// TIA Portal project "uppgift2IndustriellIT" (V18)

(* hardware
DEVICE "S7-1500/ET200MP station_1"  S7-1500 station
   slot 0: "Rail_0"  Rack  6ES7 590-1***0-0AA0
   slot 1: "PLC_1"  CPU 1518-4 PN/DP  6ES7 518-4AP00-0AB0  V3.0
      slot 3: "CPU display_1"  6ES7591-1BA00-0AA0
      slot 32768: "PROFINET interface_1"  X1
         slot 32769: "Port_1"  X1 P1
         slot 32770: "Port_2"  X1 P2
      slot 33024: "PROFINET interface_2"  X2
         slot 33025: "Port_1"  X2 P1
      slot 33280: "PROFINET interface GBIT_3"  X3
         slot 33281: "Port_1"  X3 P1
      slot 33536: "DP interface_1"  X4
      slot 34817: "Virtual CP interface port_1"  Virtual CP interface port  Virtual CP interface port
DEVICE "HMI_1"  KTP700 Mobile
   slot 0: "HMI_1"  KTP700 Mobile  6AV2 125-2GB03-0AX0  17.0.0.0
   slot 1: "HMI_RT_1"  KTP700 Mobile  6AV2 125-2GB03-0AX0  17.0.0.0
   slot 5: "HMI_1.IE_CP_1"  PROFINET Interface  17.0.0.0
      slot 1: "PROFINET Interface_1"  PROFINET Interface
         slot 1: "Port_1"  Port
DEVICE "PC-System_1"  SIMATIC PC station
   slot 0: "SIMATIC PC station"  Rail  SIMATIC PC-Station  V1.0
      slot 125: "Stationmanager"  Station_Manager  V6.0.4
   slot 1: "HMI_RT_2"  WinCC RT Advanced  6AV2 104-0xxxx-xxxx  17.0.0.0
      slot 33792: "Computer interface"  Host interface
   slot 2: "IE general_1"  IE General  IE_CP  V8.2.0
      slot 1: "PROFINET interface"  IEGeneral.Interface.8.2.0
*)

// ===== PLC "PLC_1"  CPU 1518-4 PN/DP =====

VAR_GLOBAL   // PLC tag table "Clock/Flanks"
   "Clock_Byte" AT %MB0 : Byte;
   "Clock_10Hz" AT %M0.0 : Bool;
   "Clock_5Hz" AT %M0.1 : Bool;
   "Clock_2.5Hz" AT %M0.2 : Bool;
   "Clock_2Hz" AT %M0.3 : Bool;
   "Clock_1.25Hz" AT %M0.4 : Bool;
   "Clock_1Hz" AT %M0.5 : Bool;
   "Clock_0.625Hz" AT %M0.6 : Bool;
   "Clock_0.5Hz" AT %M0.7 : Bool;
   "PartExitFlank" AT %I3.0 : Bool;
   "CraneExitPosFlank" AT %I3.1 : Bool;
   "HmiEntryFlank" AT %I4.0 : Bool;
   "HmiFlankExit" AT %I4.1 : Bool;
   "FoundToUnloadFlank" AT %I4.2 : Bool;
   "HmiFlankLoad" AT %I5.0 : Bool;
   "HmiFlankUnload" AT %I5.2 : Bool;
   "VisionErrorFlank" AT %I5.4 : Bool;
END_VAR

VAR_GLOBAL   // PLC tag table "FactoryIO"
   "Start Button" AT %I0.0 : Bool;
   "Reset Button" AT %I0.1 : Bool;
   "Stop Button (NC)" AT %I0.2 : Bool;
   "Emergency Stop (NC)" AT %I0.3 : Bool;
   "Part At Entry (NC)" AT %I0.4 : Bool;
   "Part At Load (NC)" AT %I0.5 : Bool;
   "Part At Unload (NC)" AT %I0.6 : Bool;
   "Part At Exit (NC)" AT %I0.7 : Bool;
   "Crane is at Entry-Pos" AT %I1.0 : Bool;
   "Crane is at Exit-Pos" AT %I1.1 : Bool;
   "Crane is at Default-Pos" AT %I1.2 : Bool;
   "Start Light" AT %Q0.0 : Bool;
   "Reset Light" AT %Q0.1 : Bool;
   "Stop Light" AT %Q0.2 : Bool;
   "Protection Stoplight" AT %Q0.3 : Bool;
   "Emitter" AT %Q0.4 : Bool;
   "Signal Tower Green" AT %Q0.5 : Bool;
   "Signal Tower Yellow" AT %Q0.6 : Bool;
   "Signal Tower Red" AT %Q0.7 : Bool;
   "Extend Crane Entry-Side" AT %Q1.0 : Bool;
   "Extend Crane Exit-Side" AT %Q1.1 : Bool;
   "Vision Sensor Entry" AT %IW24 : Int;
   "Crane Current X Position" AT %IW26 : Int;
   "Crane Current Z Position" AT %IW28 : Int;
   "Entry Conveyor" AT %QW20 : Int;
   "Loading Conveyor" AT %QW22 : Int;
   "Unloading Conveyor" AT %QW24 : Int;
   "Set Crane X Position" AT %QW26 : Int;
   "Set Crane Z Position" AT %QW28 : Int;
   "Free Slots in Storage" AT %QW30 : Int;
   "factoryiorunning" AT %I1.3 : Bool;
   "Exit conveyor" AT %QW32 : Int;
   "alarmStuck" AT %QW34 : Int;
   "alarmLoaderFull" AT %QW36 : Int;
   "alarmUnloaderEmpty" AT %QW38 : Int;
END_VAR

// folder: Databases/HmiRelated

DATA_BLOCK "HmiDb"   // DB16
{ S7_Optimized_Access := 'TRUE' }
VERSION : 0.1
   VAR
      HmiOrderMode : Struct
         HmiOrderAmount : Int;
         HmiExecuteOrder : Bool;
         HmiColorSelected : Int;
         HmiPauseOrder : Bool;
         OrderDelivered : Int;
      END_STRUCT;
      ActivateAcutator : Struct
         HmiRunEntryConv : Bool;
         HmiRunExitConv : Bool;
         HmiExtendEntry : Bool;
         HmiExtendExit : Bool;
         HmiRunLoadConv : Bool;
         HmiRunUnloadConv : Bool;
         hmilighttest : Bool;
      END_STRUCT;
      HmiModes : Struct
         ActivateUnloadHmi : Bool;
         HmiStopmode : Bool;
         HmiRunMode : Bool;
         HmiResetMode : Bool;
      END_STRUCT;
      BoxyMover : Int;
      BoxyMover2 : Int;
      ClearStock : Bool;
      ClearCounter : Bool;
      HmiSaveArmCalX : Bool;
      HmiSaveArmCalY : Bool;
      XListColumn : Int;
      YListColumn : Int;
      CalInputVal : Int;
      CurrentPositionX : Int;
      CurrentPositionY : Int;
      oke : String := 'yes';
   END_VAR
BEGIN
END_DATA_BLOCK

DATA_BLOCK "jogmodeDB"   // DB18
{ S7_Optimized_Access := 'TRUE' }
VERSION : 0.1
   VAR
      CraneXjog : Int;
      CraneYjog : Int;
   END_VAR
BEGIN
END_DATA_BLOCK

// folder: Databases/SCLdb

DATA_BLOCK "PositionArray"   // DB9
{ S7_Optimized_Access := 'TRUE' }
VERSION : 0.1
   VAR RETAIN
      YposCraneMM : Array[0..5] of Int;
      XposCraneMM : Array[0..8] of Int;
   END_VAR
BEGIN
   YposCraneMM[0] := 380;
   YposCraneMM[1] := 1540;
   YposCraneMM[2] := 2680;
   YposCraneMM[3] := 3820;
   YposCraneMM[4] := 4950;
   YposCraneMM[5] := 6000;
   XposCraneMM[0] := 1490;
   XposCraneMM[1] := 2635;
   XposCraneMM[2] := 3750;
   XposCraneMM[3] := 4860;
   XposCraneMM[4] := 6000;
   XposCraneMM[5] := 7145;
   XposCraneMM[6] := 8260;
   XposCraneMM[7] := 9380;
   XposCraneMM[8] := 10500;
END_DATA_BLOCK

DATA_BLOCK "PositionUnload_DB"   // DB10
{ S7_Optimized_Access := 'TRUE' }
VERSION : 0.1
// stored: InstanceOfName PositionUnload
"PositionUnload"
BEGIN
END_DATA_BLOCK

DATA_BLOCK "AlreadyFilledSlotArray"   // DB11
{ S7_Optimized_Access := 'TRUE' }
VERSION : 0.1
   VAR RETAIN
      Row1Y : Array[0..5] of Int;   // siffran i array namnet indikterar X axeln: T.ex. Row3Y visar om column 3 är fylld med lådor och index siffran i arrayn indikerar vilken våning i columen som är fylld
      Row2Y : Array[0..5] of Int;
      Row3Y : Array[0..5] of Int;
      Row4Y : Array[0..5] of Int;
      Row5Y : Array[0..5] of Int;
      Row6Y : Array[0..5] of Int;
      Row7Y : Array[0..5] of Int;
      Row8Y : Array[0..5] of Int;
      Row9Y : Array[0..5] of Int;
   END_VAR
BEGIN
   Row4Y[5] := 0;
   Row4Y[4] := 0;
   Row4Y[3] := 0;
   Row4Y[2] := 0;
   Row4Y[1] := 0;
   Row4Y[0] := 0;
   Row3Y[0] := 0;
   Row3Y[1] := 0;
   Row3Y[2] := 0;
   Row3Y[3] := 0;
   Row3Y[4] := 0;
   Row3Y[5] := 0;
   Row2Y[5] := 0;
   Row2Y[4] := 0;
   Row2Y[3] := 0;
   Row2Y[2] := 0;
   Row2Y[1] := 0;
   Row2Y[0] := 0;
   Row8Y[5] := 0;
   Row8Y[4] := 0;
   Row8Y[3] := 0;
   Row8Y[2] := 0;
   Row8Y[1] := 0;
   Row8Y[0] := 0;
   Row7Y[5] := 0;
   Row7Y[4] := 0;
   Row1Y[5] := 0;
   Row1Y[4] := 0;
   Row1Y[3] := 0;
   Row1Y[2] := 0;
   Row1Y[1] := 0;
   Row1Y[0] := 0;
   Row9Y[5] := 0;
   Row9Y[4] := 0;
   Row9Y[3] := 0;
   Row9Y[2] := 0;
   Row9Y[1] := 0;
   Row9Y[0] := 0;
   Row5Y[5] := 0;
   Row5Y[4] := 0;
   Row5Y[3] := 0;
   Row5Y[2] := 0;
   Row5Y[1] := 0;
   Row5Y[0] := 0;
   Row6Y[5] := 0;
   Row6Y[4] := 0;
   Row6Y[3] := 0;
   Row6Y[2] := 0;
   Row6Y[1] := 0;
   Row6Y[0] := 0;
   Row7Y[3] := 0;
   Row7Y[2] := 0;
   Row7Y[1] := 0;
   Row7Y[0] := 0;
END_DATA_BLOCK

DATA_BLOCK "PositionsLOAD_DB"   // DB13
{ S7_Optimized_Access := 'TRUE' }
VERSION : 0.1
// stored: InstanceOfName PositionsLoad
"PositionsLoad"
BEGIN
END_DATA_BLOCK

DATA_BLOCK "resetFill_DB"   // DB21
{ S7_Optimized_Access := 'TRUE' }
VERSION : 0.1
// stored: InstanceOfName resetFill
"resetFill"
BEGIN
END_DATA_BLOCK

// folder: Databases/input/outputDB

DATA_BLOCK "InputsDB"   // DB1
{ S7_Optimized_Access := 'TRUE' }
VERSION : 0.1
   VAR RETAIN
      ConvertedConveyors : Struct
         EntryConvSensorVal : Int := 7500;
         LoadingConvSensorVal : Int := 7500;
         EntryConvScalex : Real;
         LoadingConvScalex : Real;
         ExitConvSensorVal : Int := 7500;
         ExitConvScaleX : Real;
         UnloadingScaleX : Real;
         UnloadingSensorVal : Int := 7500;
      END_STRUCT;
   END_VAR
   VAR
      ConveyorSaveCalVal : Struct
         Normxconverter : Real;
         Save : Bool;
         "DisplayMm/s" : Real;
         Min : Struct
            EntryMin : Int;
            ExitMin : Int;
            LoadMin : Int;
            UnloadMin : Int;
            HmiDisplayMin : Int;
            ActualdisplayMin : Int;
         END_STRUCT;
         Max : Struct
            EntryMax : Int;
            ExitMax : Int;
            LoadMax : Int;
            UnloadMax : Int;
            HmiDisplayMax : Int;
            ActualdisplayMax : Int;
         END_STRUCT;
      END_STRUCT;
      RunConveyor : Struct
         RunEntryConveyor : Bool;
         RunLoadingConveyor : Bool;
         RunUnloadingConveyor : Bool;
         RunExitConveyor : Bool;
      END_STRUCT;
      Crane : Struct
         X : Struct
            XSensorValueNormx : Real;
            XSensorValueScaleX : Int;
            SaveX : Int;
         END_STRUCT;
         Y : Struct
            YSensorValueNormx : Real;
            YSensorValueScalex : Int;
            SaveY : Int;
         END_STRUCT;
         RunArmX : Bool;
         RunArmY : Bool;
      END_STRUCT;
      Sensors : Struct
         "Part Entry" : Bool;
         "Part Load" : Bool;
         "Part Unload" : Bool;
         "Part Exit" : Bool;
         "Crane Entry" : Bool;
         "Crane Exit" : Bool;
         "Crane Default" : Bool;
         "Color Sensor" : Int;
      END_STRUCT;
      Conditions : Struct
         ProtectedStop : Bool;
         HasBeenJogging : Bool;
         VisionError : Bool;
      END_STRUCT;
      FreeSlotCounter : Int := 54;
      ErrorStuck : Bool;
      ConveyorCalibrationPicker : Int := 10;   // Slidern i hmin
      ConveyorCalibrationBarSlider : Int := 7500;
      ConveyorCalibrationBarSliderTEMP : Int;
      YisMoving : Bool;
      XisMoving : Bool;   // Används endast för hmin just nu
      Math200 : Int := 200;
      Math10 : Int;
      AdjustX : Int;
      AdjustY : Int;
      PressAdjustX : Bool;
      PressAdjustY : Bool;
      totalcounter : Int;
      totalremovedcounter : Int;
   END_VAR
BEGIN
END_DATA_BLOCK

DATA_BLOCK "OutputsDB"   // DB2
{ S7_Optimized_Access := 'TRUE' }
VERSION : 0.1
   VAR
      CraneOutput : Struct
         Xmm : Int;
         Xnormx : Real;
         XScalex : Int;
         Ymm : Int;
         Ynormx : Real;
         YScalex : Int;
      END_STRUCT;
      ForkController : Struct
         MoveForkExitLoad : Bool;
         MoveForkEntryLoad : Bool;
         SafetyStopExitUnload : Bool;
      END_STRUCT;
   END_VAR
BEGIN
END_DATA_BLOCK

DATA_BLOCK "Modes"   // DB3
{ S7_Optimized_Access := 'TRUE' }
VERSION : 0.1
   VAR
      Modes : Struct
         RunMode : Bool;
         ResetMode : Bool;
         Unloadmode : Bool;
         RunUnloadConveyor : Bool;
         StoppestMode : Bool;
         JogMode : Bool;
         OrderMode : Bool;
      END_STRUCT;
      Sequences : Struct
         SequenceLoader : Int := 10;
         SequenceUnloader : Int := 10;
         ResetModeSequence : Int := 10;
         SafetyStopSequence : Int := 10;
      END_STRUCT;
      StopMethods : Struct
         SafetyStop : Bool;
         ProductionStop : Bool := true;
      END_STRUCT;
   END_VAR
BEGIN
END_DATA_BLOCK

DATA_BLOCK "ColorDB"   // DB5
{ S7_Optimized_Access := 'TRUE' }
VERSION : 0.1
   VAR
      Gray : Int;
      Green : Int;
      Blue : Int;
      isGray : Int := 1;
      isBlue : Int := 2;
      isGreen : Int := 3;
   END_VAR
BEGIN
END_DATA_BLOCK

// folder: System blocks/Program resources

DATA_BLOCK "ResetWaiterTimer"   // DB4
{ S7_Optimized_Access := 'TRUE' }
AUTHOR : Simatic
FAMILY : IEC
NAME : IEC_TMR
VERSION : 1.0
// stored: InstanceOfName IEC_TIMER
"IEC_TIMER"
BEGIN
END_DATA_BLOCK

DATA_BLOCK "ColorCounter1"   // DB6
{ S7_Optimized_Access := 'TRUE' }
AUTHOR : Simatic
FAMILY : IEC
NAME : CNTR
VERSION : 1.0
// stored: InstanceOfName IEC_COUNTER
"IEC_COUNTER"
BEGIN
END_DATA_BLOCK

DATA_BLOCK "ColorCouter2"   // DB7
{ S7_Optimized_Access := 'TRUE' }
AUTHOR : Simatic
FAMILY : IEC
NAME : CNTR
VERSION : 1.0
// stored: InstanceOfName IEC_COUNTER
"IEC_COUNTER"
BEGIN
END_DATA_BLOCK

DATA_BLOCK "ColorCounter3"   // DB8
{ S7_Optimized_Access := 'TRUE' }
AUTHOR : Simatic
FAMILY : IEC
NAME : CNTR
VERSION : 1.0
// stored: InstanceOfName IEC_COUNTER
"IEC_COUNTER"
BEGIN
END_DATA_BLOCK

DATA_BLOCK "SclDelay"   // DB12
{ S7_Optimized_Access := 'TRUE' }
AUTHOR : Simatic
FAMILY : IEC
NAME : IEC_TMR
VERSION : 1.0
// stored: InstanceOfName IEC_TIMER
"IEC_TIMER"
BEGIN
END_DATA_BLOCK

DATA_BLOCK "SclDelay2"   // DB14
{ S7_Optimized_Access := 'TRUE' }
AUTHOR : Simatic
FAMILY : IEC
NAME : IEC_TMR
VERSION : 1.0
// stored: InstanceOfName IEC_TIMER
"IEC_TIMER"
BEGIN
END_DATA_BLOCK

DATA_BLOCK "ForkWaiter"   // DB15
{ S7_Optimized_Access := 'TRUE' }
AUTHOR : Simatic
FAMILY : IEC
NAME : IEC_TMR
VERSION : 1.0
// stored: InstanceOfName IEC_TIMER
"IEC_TIMER"
BEGIN
END_DATA_BLOCK

DATA_BLOCK "StuckTimer"   // DB17
{ S7_Optimized_Access := 'TRUE' }
AUTHOR : Simatic
FAMILY : IEC
NAME : IEC_TMR
VERSION : 1.0
// stored: InstanceOfName IEC_TIMER
"IEC_TIMER"
BEGIN
END_DATA_BLOCK

DATA_BLOCK "FreeSlotCounter"   // DB19
{ S7_Optimized_Access := 'TRUE' }
AUTHOR : Simatic
FAMILY : IEC
NAME : CNTR
VERSION : 1.0
// stored: InstanceOfName IEC_COUNTER
"IEC_COUNTER"
BEGIN
   CV := 54;
END_DATA_BLOCK

DATA_BLOCK "OrderDeliverCounter"   // DB20
{ S7_Optimized_Access := 'TRUE' }
AUTHOR : Simatic
FAMILY : IEC
NAME : CNTR
VERSION : 1.0
// stored: InstanceOfName IEC_COUNTER
"IEC_COUNTER"
BEGIN
END_DATA_BLOCK

DATA_BLOCK "totalcounter"   // DB22
{ S7_Optimized_Access := 'TRUE' }
AUTHOR : Simatic
FAMILY : IEC
NAME : CNTR
VERSION : 1.0
// stored: InstanceOfName IEC_COUNTER
"IEC_COUNTER"
BEGIN
END_DATA_BLOCK

DATA_BLOCK "totalcounterremoved"   // DB23
{ S7_Optimized_Access := 'TRUE' }
AUTHOR : Simatic
FAMILY : IEC
NAME : CNTR
VERSION : 1.0
// stored: InstanceOfName IEC_COUNTER
"IEC_COUNTER"
BEGIN
END_DATA_BLOCK

DATA_BLOCK "ResetWaiterTimer2"   // DB24
{ S7_Optimized_Access := 'TRUE' }
AUTHOR : Simatic
FAMILY : IEC
NAME : IEC_TMR
VERSION : 1.0
// stored: InstanceOfName IEC_TIMER
"IEC_TIMER"
BEGIN
END_DATA_BLOCK

DATA_BLOCK "waittimer3"   // DB25
{ S7_Optimized_Access := 'TRUE' }
AUTHOR : Simatic
FAMILY : IEC
NAME : IEC_TMR
VERSION : 1.0
// stored: InstanceOfName IEC_TIMER
"IEC_TIMER"
BEGIN
END_DATA_BLOCK

// folder: (top level)

ORGANIZATION_BLOCK "Main"   // OB1, LAD, ProgramCycle
TITLE = "Main Program Sweep (Cycle)"
{ S7_Optimized_Access := 'TRUE' }
VERSION : 0.1
   VAR_INPUT
      Initial_Call : Bool;   // Initial call of this OB
      Remanence : Bool;   // =True, if remanent data are available
   END_VAR
BEGIN

REGION Network 1
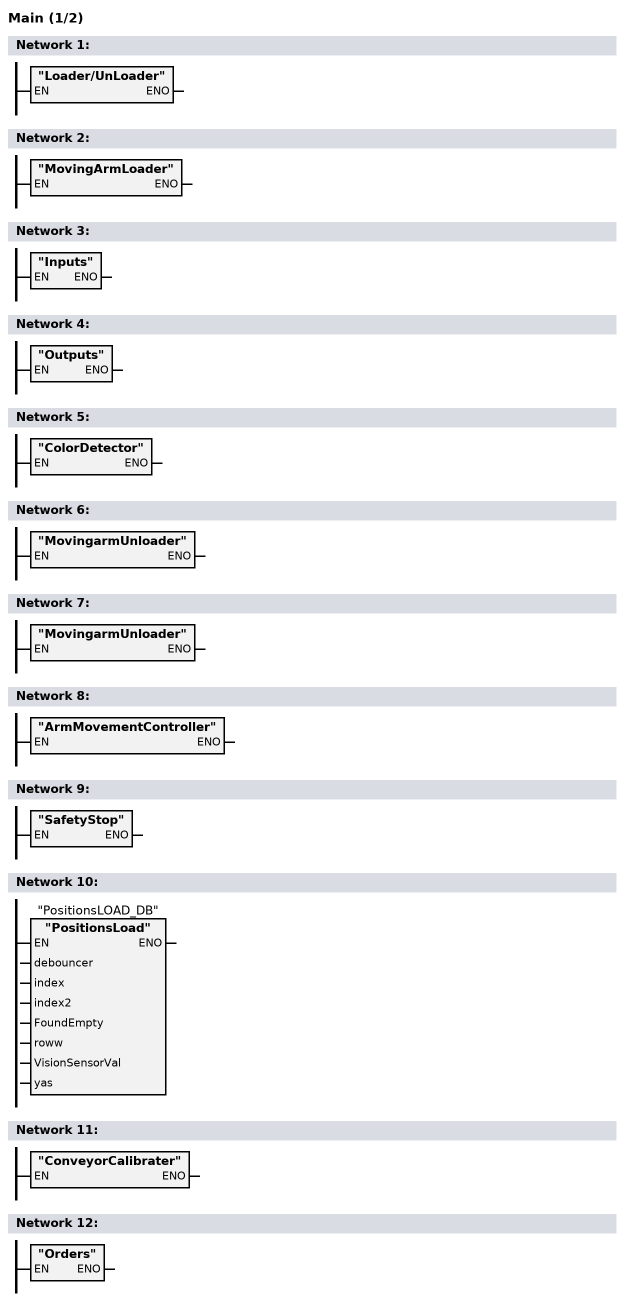
   RUNG wire#powerrail
      "Loader/UnLoader"()
   END_RUNG
   // the same network as SCL:
   "Loader/UnLoader"();
END_REGION

REGION Network 2
   RUNG wire#powerrail
      "MovingArmLoader"()
   END_RUNG
   // the same network as SCL:
   "MovingArmLoader"();
END_REGION

REGION Network 3
   RUNG wire#powerrail
      "Inputs"()
   END_RUNG
   // the same network as SCL:
   "Inputs"();
END_REGION

REGION Network 4
   RUNG wire#powerrail
      "Outputs"()
   END_RUNG
   // the same network as SCL:
   "Outputs"();
END_REGION

REGION Network 5
   RUNG wire#powerrail
      "ColorDetector"()
   END_RUNG
   // the same network as SCL:
   "ColorDetector"();
END_REGION

REGION Network 6
   RUNG wire#powerrail
      "MovingarmUnloader"()
   END_RUNG
   // the same network as SCL:
   "MovingarmUnloader"();
END_REGION

REGION Network 7
   RUNG wire#powerrail
      "MovingarmUnloader"()
   END_RUNG
   // the same network as SCL:
   "MovingarmUnloader"();
END_REGION

REGION Network 8
   RUNG wire#powerrail
      "ArmMovementController"()
   END_RUNG
   // the same network as SCL:
   "ArmMovementController"();
END_REGION

REGION Network 9
   RUNG wire#powerrail
      "SafetyStop"()
   END_RUNG
   // the same network as SCL:
   "SafetyStop"();
END_REGION

REGION Network 10
   RUNG wire#powerrail
      "PositionsLOAD_DB"(debouncer :=, index :=, index2 :=, FoundEmpty :=, roww :=, VisionSensorVal :=, yas :=)
   END_RUNG
   // the same network as SCL:
   "PositionsLOAD_DB"();   // "PositionsLoad"
END_REGION

REGION Network 11
   RUNG wire#powerrail
      "ConveyorCalibrater"()
   END_RUNG
   // the same network as SCL:
   "ConveyorCalibrater"();
END_REGION

REGION Network 12
   RUNG wire#powerrail
      "Orders"()
   END_RUNG
   // the same network as SCL:
   "Orders"();
END_REGION

REGION Network 13
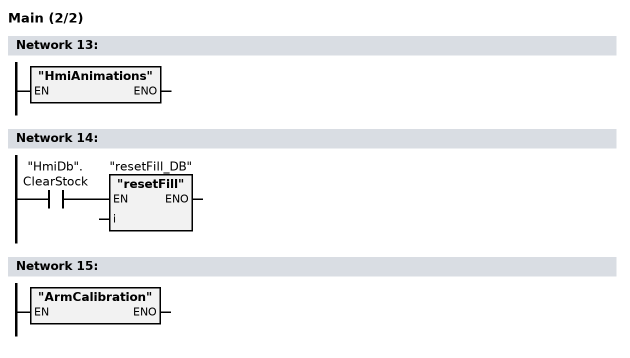
   RUNG wire#powerrail
      "HmiAnimations"()
   END_RUNG
   // the same network as SCL:
   "HmiAnimations"();
END_REGION

REGION Network 14
   RUNG wire#powerrail
      Contact( "HmiDb".ClearStock )
      "resetFill_DB"(i :=)
   END_RUNG
   // the same network as SCL:
   IF "HmiDb".ClearStock THEN
       "resetFill_DB"();   // "resetFill"
   END_IF;
END_REGION

REGION Network 15
   RUNG wire#powerrail
      "ArmCalibration"()
   END_RUNG
   // the same network as SCL:
   "ArmCalibration"();
END_REGION
END_ORGANIZATION_BLOCK

// folder: Functions/ArmGroup

FUNCTION "Loader/UnLoader" : Void   // FC1, LAD
{ S7_Optimized_Access := 'TRUE' }
VERSION : 0.1
   VAR_TEMP   // added for the SCL form of the ladder/FBD networks
      _w1 : Bool;
      _w2 : Bool;
   END_VAR
BEGIN

REGION Network 1: Om på sekvens 1 då kör emittern
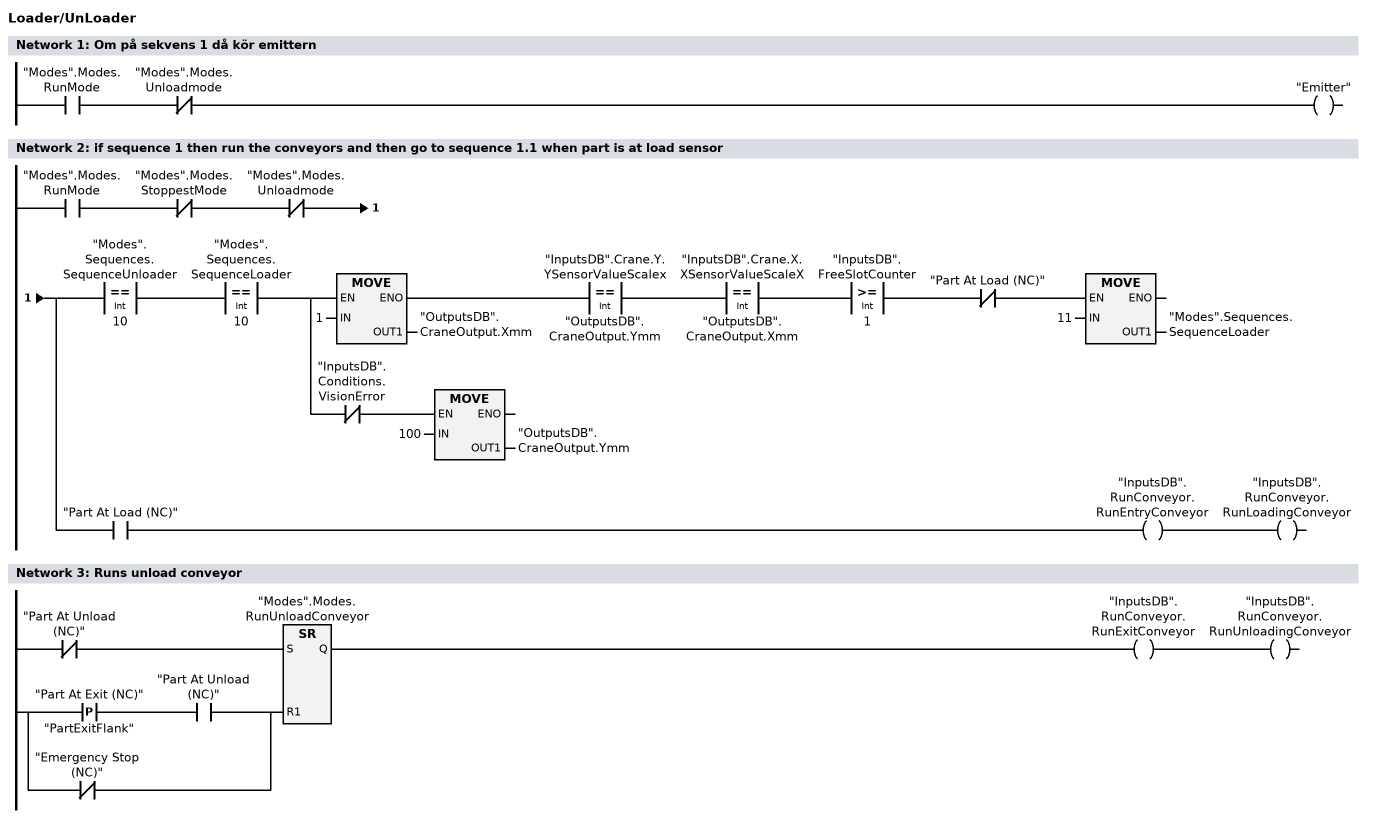
   RUNG wire#powerrail
      Contact( "Modes".Modes.RunMode )
      I_Contact( "Modes".Modes.Unloadmode )
      Coil( "Emitter" )
   END_RUNG
   // the same network as SCL:
   "Emitter" := "Modes".Modes.RunMode AND NOT "Modes".Modes.Unloadmode;
END_REGION

REGION Network 2: if sequence 1 then run the conveyors and then go to sequence 1.1 when part is at load sensor
   RUNG wire#powerrail
      Contact( "Modes".Modes.RunMode )
      I_Contact( "Modes".Modes.StoppestMode )
      I_Contact( "Modes".Modes.Unloadmode )
      wire#w1
      { S7_Templates := "SrcType := Int" } EQ_Contact(in1 := "Modes".Sequences.SequenceUnloader, in2 := 10)
      { S7_Templates := "SrcType := Int" } EQ_Contact(in1 := "Modes".Sequences.SequenceLoader, in2 := 10)
      wire#w2
      Move(in := 1, out1 => "OutputsDB".CraneOutput.Xmm)
      { S7_Templates := "SrcType := Int" } EQ_Contact(in1 := "InputsDB".Crane.Y.YSensorValueScalex, in2 := "OutputsDB".CraneOutput.Ymm)
      { S7_Templates := "SrcType := Int" } EQ_Contact(in1 := "InputsDB".Crane.X.XSensorValueScaleX, in2 := "OutputsDB".CraneOutput.Xmm)
      { S7_Templates := "SrcType := Int" } GE_Contact(in1 := "InputsDB".FreeSlotCounter, in2 := 1)
      I_Contact( "Part At Load (NC)" )
      Move(in := 11, out1 => "Modes".Sequences.SequenceLoader)
   END_RUNG
   RUNG wire#w2
      I_Contact( "InputsDB".Conditions.VisionError )
      Move(in := 100, out1 => "OutputsDB".CraneOutput.Ymm)
   END_RUNG
   RUNG wire#w1
      Contact( "Part At Load (NC)" )
      Coil( "InputsDB".RunConveyor.RunEntryConveyor )
      Coil( "InputsDB".RunConveyor.RunLoadingConveyor )
   END_RUNG
   // the same network as SCL:
   #_w1 := "Modes".Modes.RunMode AND NOT "Modes".Modes.StoppestMode AND NOT "Modes".Modes.Unloadmode;
   #_w2 := #_w1 AND ("Modes".Sequences.SequenceUnloader = 10) AND ("Modes".Sequences.SequenceLoader = 10);
   IF #_w2 THEN "OutputsDB".CraneOutput.Xmm := 1; END_IF;
   IF #_w2 AND ("InputsDB".Crane.Y.YSensorValueScalex = "OutputsDB".CraneOutput.Ymm) AND ("InputsDB".Crane.X.XSensorValueScaleX = "OutputsDB".CraneOutput.Xmm) AND ("InputsDB".FreeSlotCounter >= 1) AND NOT "Part At Load (NC)" THEN
       "Modes".Sequences.SequenceLoader := 11;
   END_IF;
   IF #_w2 AND NOT "InputsDB".Conditions.VisionError THEN "OutputsDB".CraneOutput.Ymm := 100; END_IF;
   "InputsDB".RunConveyor.RunEntryConveyor := #_w1 AND "Part At Load (NC)";
   "InputsDB".RunConveyor.RunLoadingConveyor := "InputsDB".RunConveyor.RunEntryConveyor;
END_REGION

REGION Network 3: Runs unload conveyor
   RUNG wire#powerrail
      I_Contact( "Part At Unload (NC)" )
      S_SR(operand := "Modes".Modes.RunUnloadConveyor, r1 := wire#w1)
      Coil( "InputsDB".RunConveyor.RunExitConveyor )
      Coil( "InputsDB".RunConveyor.RunUnloadingConveyor )
   END_RUNG
   RUNG wire#powerrail
      P_Contact(operand := "Part At Exit (NC)", bit := "PartExitFlank")
      Contact( "Part At Unload (NC)" )
   END_RUNG wire#w1
   RUNG wire#powerrail
      I_Contact( "Emergency Stop (NC)" )
   END_RUNG wire#w1
   // the same network as SCL:
   #_w1 := "Part At Exit (NC)" AND NOT "PartExitFlank";   // rising edge of "Part At Exit (NC)"
   "PartExitFlank" := "Part At Exit (NC)";
   IF NOT "Part At Unload (NC)" THEN
       "Modes".Modes.RunUnloadConveyor := TRUE;   // SR flip-flop
   END_IF;
   IF (#_w1 AND "Part At Unload (NC)") OR NOT "Emergency Stop (NC)" THEN
       "Modes".Modes.RunUnloadConveyor := FALSE;
   END_IF;
   "InputsDB".RunConveyor.RunExitConveyor := "Modes".Modes.RunUnloadConveyor;
   "InputsDB".RunConveyor.RunUnloadingConveyor := "Modes".Modes.RunUnloadConveyor;
END_REGION
END_FUNCTION

FUNCTION "MovingArmLoader" : Void   // FC2, FBD
{ S7_Optimized_Access := 'TRUE' }
VERSION : 0.1
   VAR_TEMP   // added for the SCL form of the ladder/FBD networks
      _w1 : Bool;
   END_VAR
BEGIN

REGION Network 1: Extend the crane and then go to next sequence
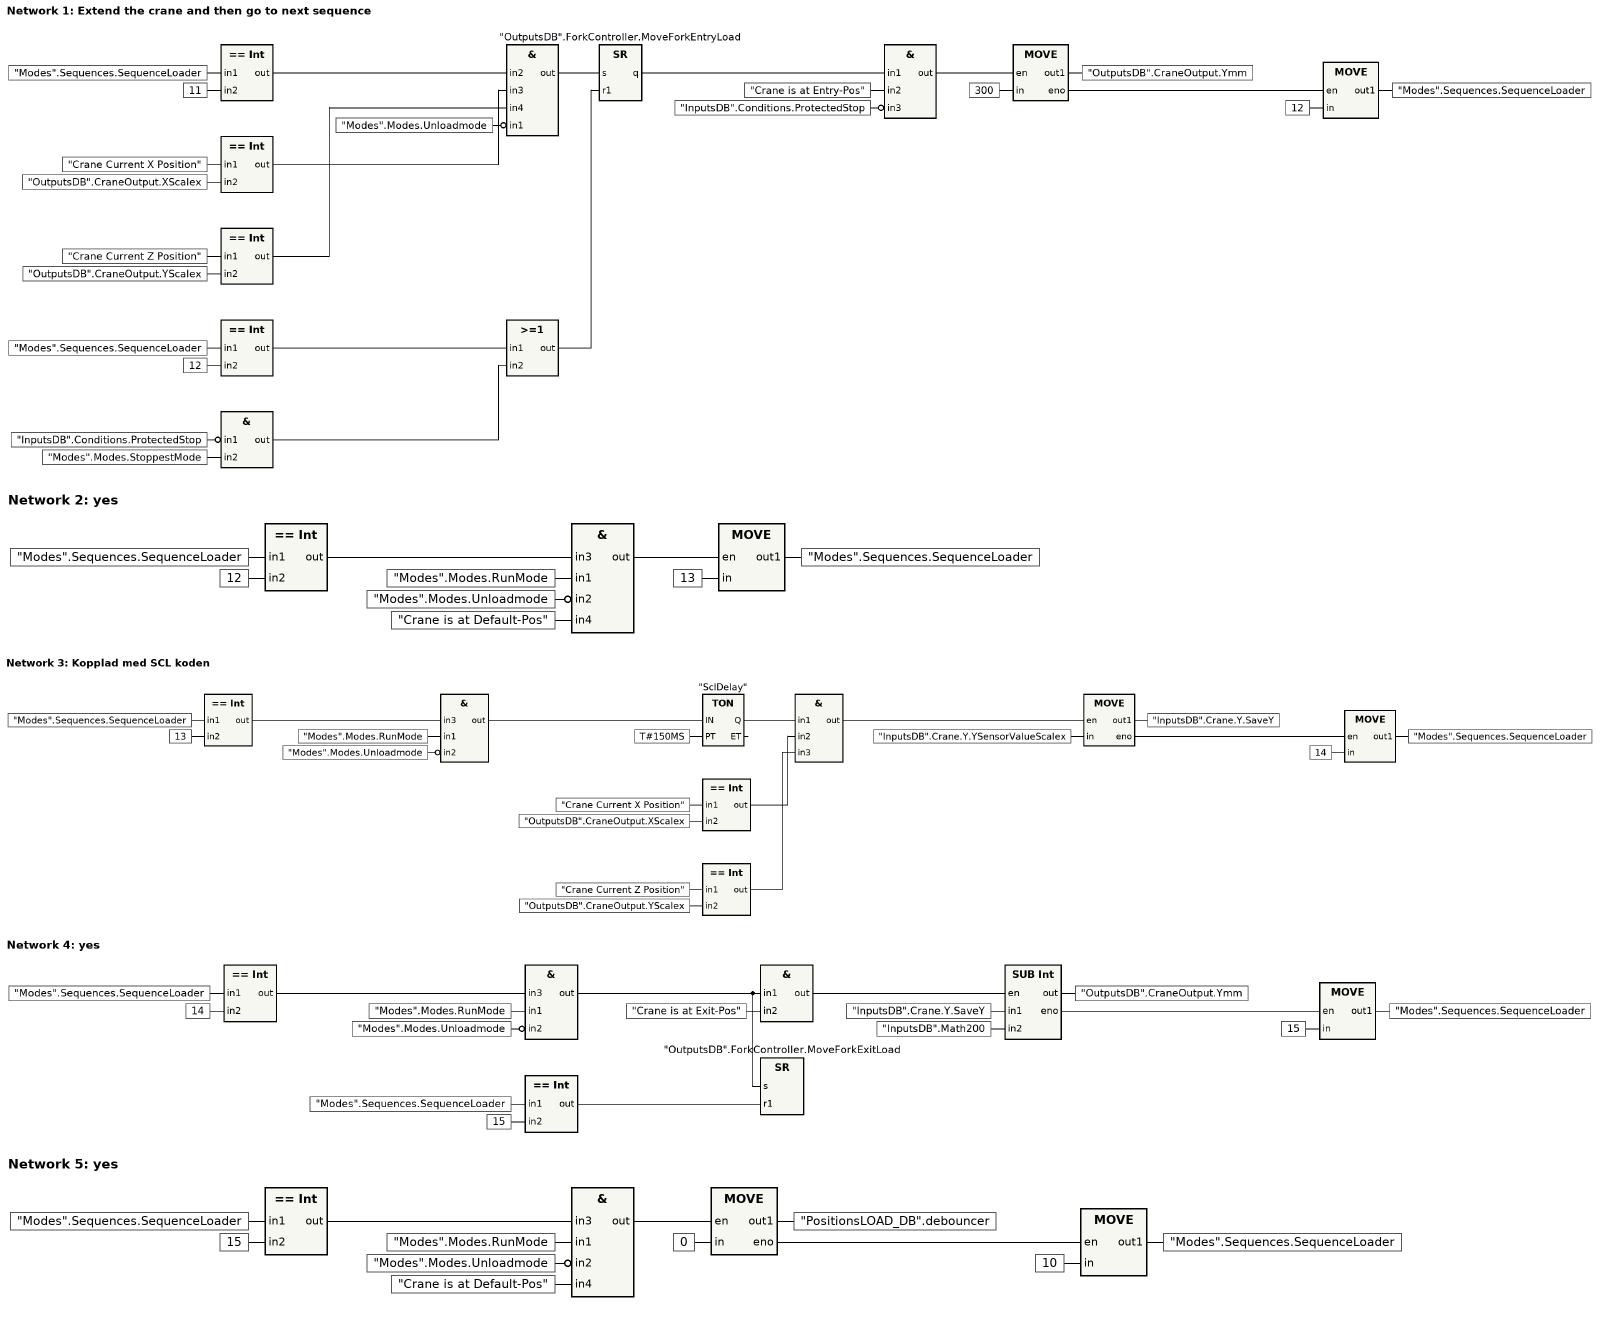
   IF ("Modes".Sequences.SequenceLoader = 11) AND ("Crane Current X Position" = "OutputsDB".CraneOutput.XScalex) AND ("Crane Current Z Position" = "OutputsDB".CraneOutput.YScalex) AND NOT "Modes".Modes.Unloadmode THEN
       "OutputsDB".ForkController.MoveForkEntryLoad := TRUE;   // SR flip-flop
   END_IF;
   IF ("Modes".Sequences.SequenceLoader = 12) OR (NOT "InputsDB".Conditions.ProtectedStop AND "Modes".Modes.StoppestMode) THEN
       "OutputsDB".ForkController.MoveForkEntryLoad := FALSE;
   END_IF;
   IF "OutputsDB".ForkController.MoveForkEntryLoad AND "Crane is at Entry-Pos" AND NOT "InputsDB".Conditions.ProtectedStop THEN
       "OutputsDB".CraneOutput.Ymm := 300;
       "Modes".Sequences.SequenceLoader := 12;
   END_IF;
END_REGION

REGION Network 2: yes
   IF ("Modes".Sequences.SequenceLoader = 12) AND "Modes".Modes.RunMode AND NOT "Modes".Modes.Unloadmode AND "Crane is at Default-Pos" THEN
       "Modes".Sequences.SequenceLoader := 13;
   END_IF;
END_REGION

REGION Network 3: Kopplad med SCL koden
   "SclDelay".TON(IN := ("Modes".Sequences.SequenceLoader = 13) AND "Modes".Modes.RunMode AND NOT "Modes".Modes.Unloadmode,
                  PT := T#150MS);
   IF "SclDelay".Q AND ("Crane Current X Position" = "OutputsDB".CraneOutput.XScalex) AND ("Crane Current Z Position" = "OutputsDB".CraneOutput.YScalex) THEN
       "InputsDB".Crane.Y.SaveY := "InputsDB".Crane.Y.YSensorValueScalex;
       "Modes".Sequences.SequenceLoader := 14;
   END_IF;
END_REGION

REGION Network 4: yes
   #_w1 := ("Modes".Sequences.SequenceLoader = 14) AND "Modes".Modes.RunMode AND NOT "Modes".Modes.Unloadmode;
   IF #_w1 AND "Crane is at Exit-Pos" THEN
       "OutputsDB".CraneOutput.Ymm := "InputsDB".Crane.Y.SaveY - "InputsDB".Math200;
       "Modes".Sequences.SequenceLoader := 15;
   END_IF;
   IF #_w1 THEN
       "OutputsDB".ForkController.MoveForkExitLoad := TRUE;   // SR flip-flop
   END_IF;
   IF "Modes".Sequences.SequenceLoader = 15 THEN
       "OutputsDB".ForkController.MoveForkExitLoad := FALSE;
   END_IF;
END_REGION

REGION Network 5: yes
   IF ("Modes".Sequences.SequenceLoader = 15) AND "Modes".Modes.RunMode AND NOT "Modes".Modes.Unloadmode AND "Crane is at Default-Pos" THEN
       "PositionsLOAD_DB".debouncer := 0;
       "Modes".Sequences.SequenceLoader := 10;
   END_IF;
END_REGION
END_FUNCTION

FUNCTION "MovingarmUnloader" : Void   // FC6, FBD
{ S7_Optimized_Access := 'TRUE' }
VERSION : 0.1
   VAR_TEMP   // added for the SCL form of the ladder/FBD networks
      _w1 : Bool;
      _w2 : Bool;
   END_VAR
BEGIN

REGION Network 1: Gets the position from array that in the scl script Seq 1
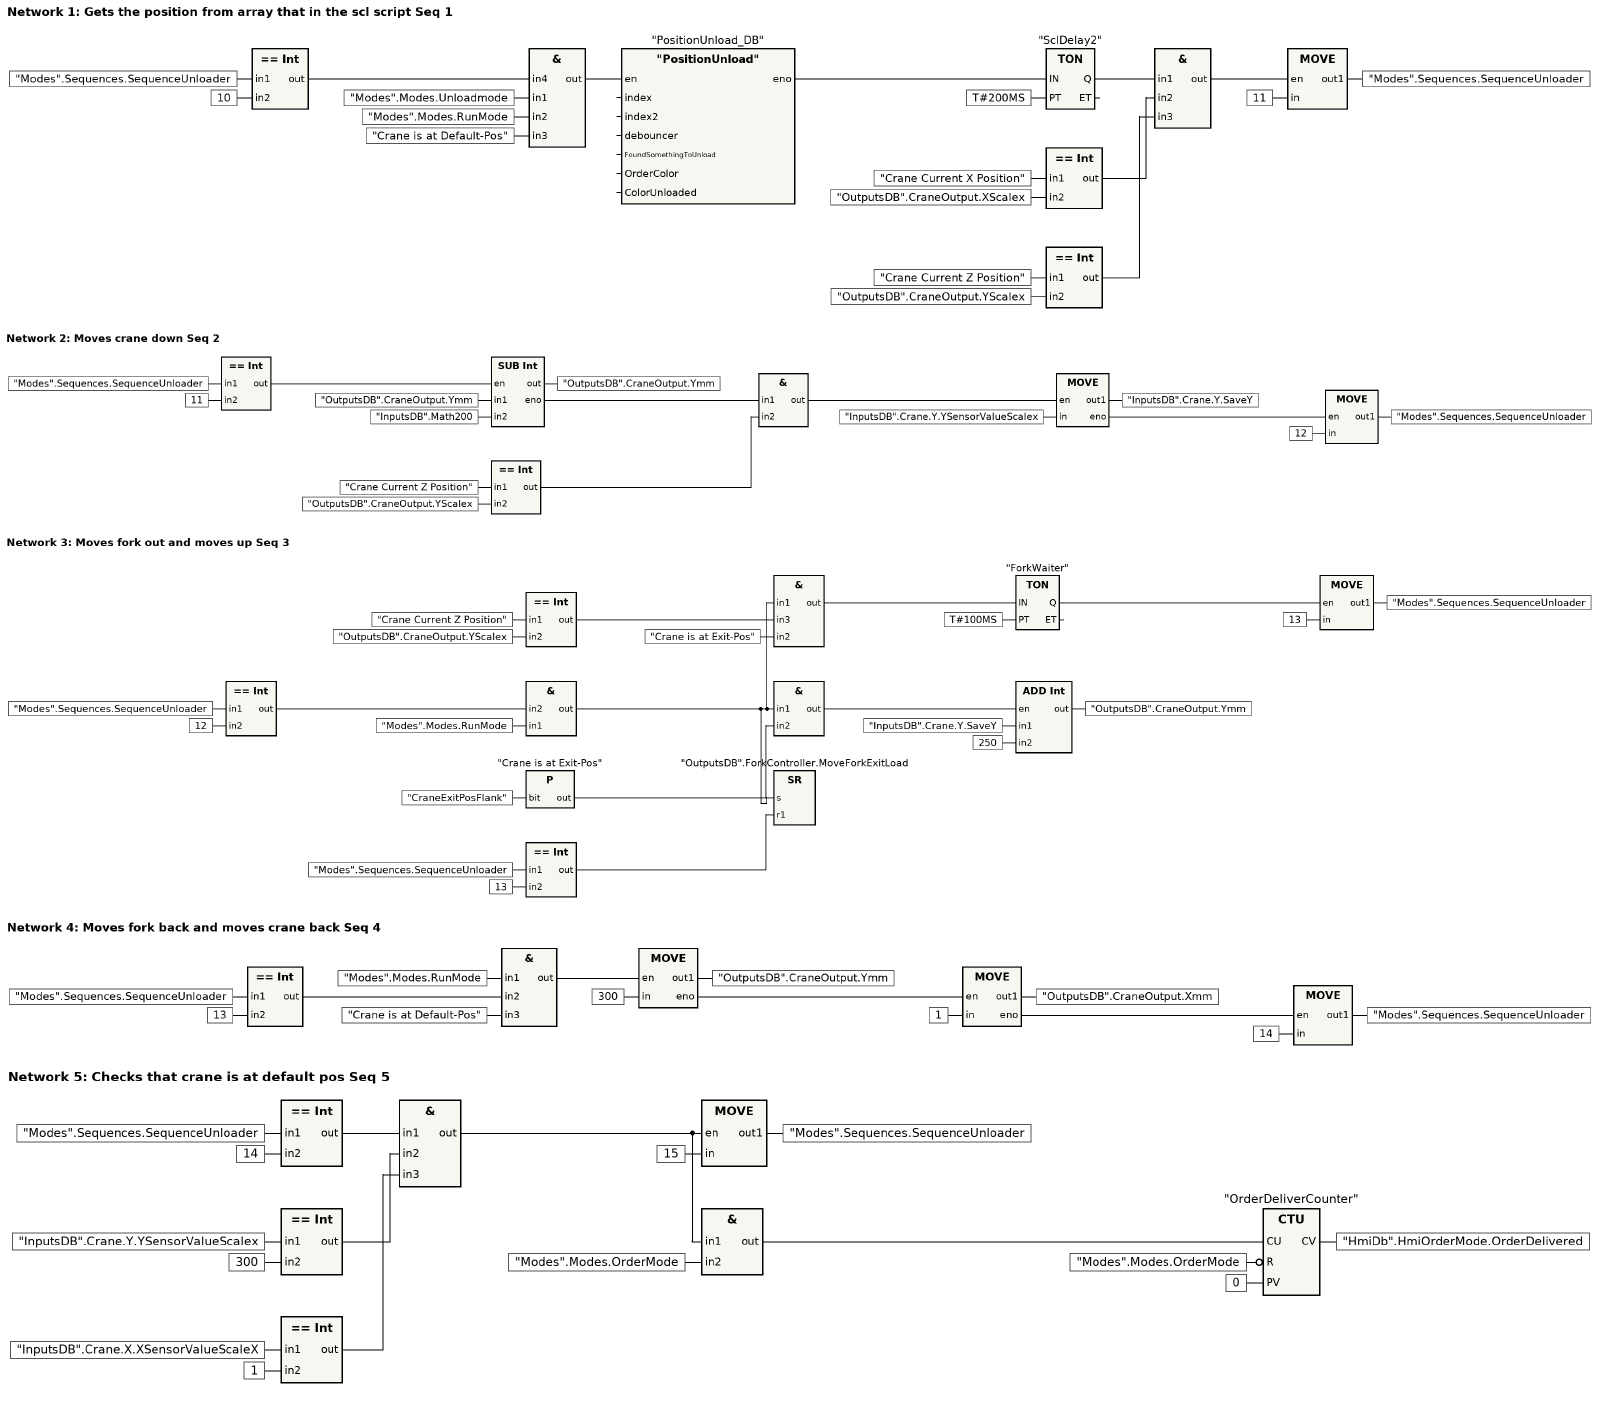
   "PositionUnload_DB"(EN := ("Modes".Sequences.SequenceUnloader = 10) AND "Modes".Modes.Unloadmode AND "Modes".Modes.RunMode AND "Crane is at Default-Pos",   // "PositionUnload"
                       ENO => #_w1);
   "SclDelay2".TON(IN := #_w1, PT := T#200MS);
   IF "SclDelay2".Q AND ("Crane Current X Position" = "OutputsDB".CraneOutput.XScalex) AND ("Crane Current Z Position" = "OutputsDB".CraneOutput.YScalex) THEN
       "Modes".Sequences.SequenceUnloader := 11;
   END_IF;
END_REGION

REGION Network 2: Moves crane down Seq 2
   #_w1 := "Modes".Sequences.SequenceUnloader = 11;
   IF #_w1 THEN "OutputsDB".CraneOutput.Ymm := "OutputsDB".CraneOutput.Ymm - "InputsDB".Math200; END_IF;
   IF #_w1 AND ("Crane Current Z Position" = "OutputsDB".CraneOutput.YScalex) THEN
       "InputsDB".Crane.Y.SaveY := "InputsDB".Crane.Y.YSensorValueScalex;
       "Modes".Sequences.SequenceUnloader := 12;
   END_IF;
END_REGION

REGION Network 3: Moves fork out and moves up Seq 3
   #_w1 := ("Modes".Sequences.SequenceUnloader = 12) AND "Modes".Modes.RunMode;
   "ForkWaiter".TON(IN := #_w1 AND ("Crane Current Z Position" = "OutputsDB".CraneOutput.YScalex) AND "Crane is at Exit-Pos",
                    PT := T#100MS);
   IF "ForkWaiter".Q THEN "Modes".Sequences.SequenceUnloader := 13; END_IF;
   #_w2 := "Crane is at Exit-Pos" AND NOT "CraneExitPosFlank";   // rising edge of "Crane is at Exit-Pos"
   "CraneExitPosFlank" := "Crane is at Exit-Pos";
   IF #_w1 AND #_w2 THEN "OutputsDB".CraneOutput.Ymm := "InputsDB".Crane.Y.SaveY + 250; END_IF;
   IF #_w1 THEN
       "OutputsDB".ForkController.MoveForkExitLoad := TRUE;   // SR flip-flop
   END_IF;
   IF "Modes".Sequences.SequenceUnloader = 13 THEN
       "OutputsDB".ForkController.MoveForkExitLoad := FALSE;
   END_IF;
END_REGION

REGION Network 4: Moves fork back and moves crane back Seq 4
   IF "Modes".Modes.RunMode AND ("Modes".Sequences.SequenceUnloader = 13) AND "Crane is at Default-Pos" THEN
       "OutputsDB".CraneOutput.Ymm := 300;
       "OutputsDB".CraneOutput.Xmm := 1;
       "Modes".Sequences.SequenceUnloader := 14;
   END_IF;
END_REGION

REGION Network 5: Checks that crane is at default pos Seq 5
   #_w1 := ("Modes".Sequences.SequenceUnloader = 14) AND ("InputsDB".Crane.Y.YSensorValueScalex = 300) AND ("InputsDB".Crane.X.XSensorValueScaleX = 1);
   IF #_w1 THEN "Modes".Sequences.SequenceUnloader := 15; END_IF;
   "OrderDeliverCounter".CTU(CU := #_w1 AND "Modes".Modes.OrderMode,
                           R := NOT "Modes".Modes.OrderMode,
                           PV := 0,
                           CV => "HmiDb".HmiOrderMode.OrderDelivered);
END_REGION

REGION Network 6: Pulls out fork Seq6
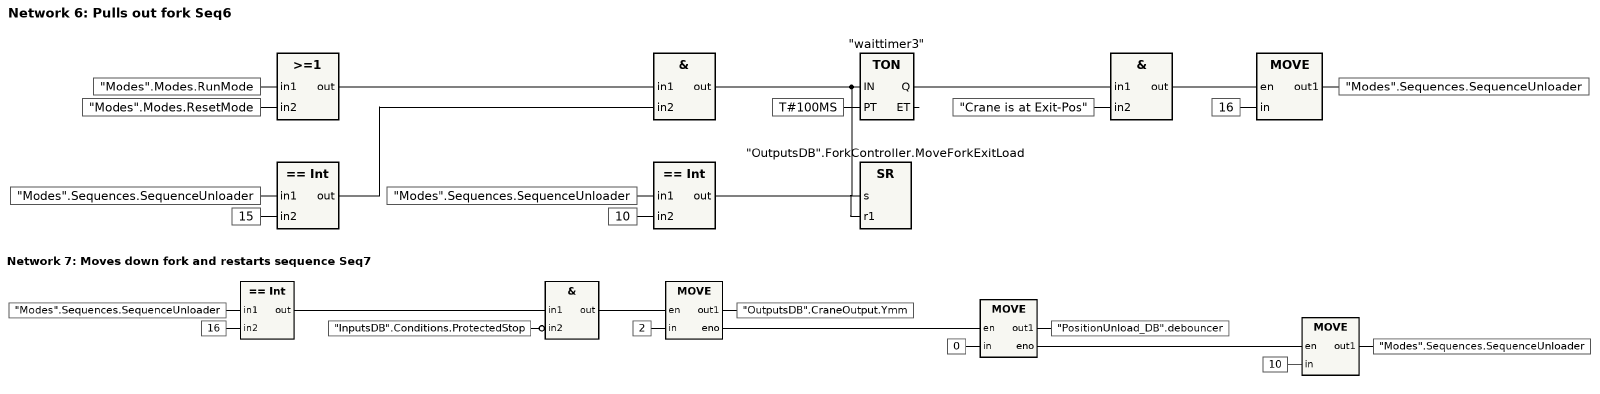
   #_w1 := ("Modes".Modes.RunMode OR "Modes".Modes.ResetMode) AND ("Modes".Sequences.SequenceUnloader = 15);
   "waittimer3".TON(IN := #_w1, PT := T#100MS);
   IF "waittimer3".Q AND "Crane is at Exit-Pos" THEN "Modes".Sequences.SequenceUnloader := 16; END_IF;
   IF #_w1 THEN
       "OutputsDB".ForkController.MoveForkExitLoad := TRUE;   // SR flip-flop
   END_IF;
   IF "Modes".Sequences.SequenceUnloader = 10 THEN
       "OutputsDB".ForkController.MoveForkExitLoad := FALSE;
   END_IF;
END_REGION

REGION Network 7: Moves down fork and restarts sequence Seq7
   IF ("Modes".Sequences.SequenceUnloader = 16) AND NOT "InputsDB".Conditions.ProtectedStop THEN
       "OutputsDB".CraneOutput.Ymm := 2;
       "PositionUnload_DB".debouncer := 0;
       "Modes".Sequences.SequenceUnloader := 10;
   END_IF;
END_REGION
END_FUNCTION

FUNCTION "ArmMovementController" : Void   // FC8, LAD
{ S7_Optimized_Access := 'TRUE' }
VERSION : 0.1
BEGIN

REGION Network 1: Controls Z(Y) axis crane and X
   // if theres a value inside "OutputsDB".CraneOutput.YScalex", thats above 1 then the arm will run
   // 
   // Example "OutputsDB".CraneOutput.YScalex" was converted from MM to sensor value
   // 
   // Example "OutputsDB".CraneOutput.Ymm" using "move" element and inputting a value in MM will then get sent, then get norm x and scalex'ed to "OutputsDB".CraneOutput.YScalex" and then move the crane